REGION Network 29: Encoder Wals Function Block
   RUNG wire#powerrail
      "FB_EncoderFeedback_Aanvoerband"(CounterTag := "EncoderBand_RawCounter", Position_Offset := "PositionManagement".Axis_1.Values."Position Offset", Pulsfactor := "PositionManagement".Axis_1.Values.Pulsfactor, Position_Correction := "PositionManagement".Axis_1.Values."Axis Correction", ReferenceRun_Command := "PositionManagement".Axis_1.Commands."Start Ref Run", ReferenceSwitch := "Zpuls_Encoder_Band", ReferencePosition := "PositionManagement".Axis_1.Values."Reference Position", Scaled_Position => #Axis1_ScaledPosition, Actual_Enc_Pos => #Axis1_ActualEncPosition, AxisDB_Connection => "PositionManagement".Data.Actual_Axis1_Position)
   END_RUNG
   // the same network as SCL:
   "FB_EncoderFeedback_Aanvoerband"(CounterTag := "EncoderBand_RawCounter",   // "FB_EncoderFeedback"
                           Position_Offset := "PositionManagement".Axis_1.Values."Position Offset",
                           Pulsfactor := "PositionManagement".Axis_1.Values.Pulsfactor,
                           Position_Correction := "PositionManagement".Axis_1.Values."Axis Correction",
                           ReferenceRun_Command := "PositionManagement".Axis_1.Commands."Start Ref Run",
                           ReferenceSwitch := "Zpuls_Encoder_Band",
                           ReferencePosition := "PositionManagement".Axis_1.Values."Reference Position",
                           Scaled_Position => #Axis1_ScaledPosition,
                           Actual_Enc_Pos => #Axis1_ActualEncPosition,
                           AxisDB_Connection => "PositionManagement".Data.Actual_Axis1_Position);
END_REGION

REGION Network 30: SystemTime
   "PLCMemory".SystemTime := TIME_TCK();
END_REGION
END_ORGANIZATION_BLOCK

// folder: Blocks

FUNCTION_BLOCK "ESB_Flash_Warning_Block"   // FB1, FBD
{ S7_Optimized_Access := 'FALSE' }
VERSION : 0.1
   VAR_INPUT
      "Safety Feedback Contact" : Bool;
      "WarningTimer Time 1" : Time := T#150ms;
      "WarningTimer Time 2" : Time := T#150ms;
   END_VAR
   VAR_OUTPUT
      "Warning Ouput Contact" : Bool;
      "ET WarningTimer 1" : Time;
      "ET WarningTimer 2" : Time;
   END_VAR
   VAR_TEMP
      SafetyTakeoverContact : Bool;
   END_VAR
   VAR_TEMP   // added for the SCL form of the ladder/FBD networks
      _w1 : Bool;
   END_VAR
BEGIN

REGION Network 1: Flash Warning
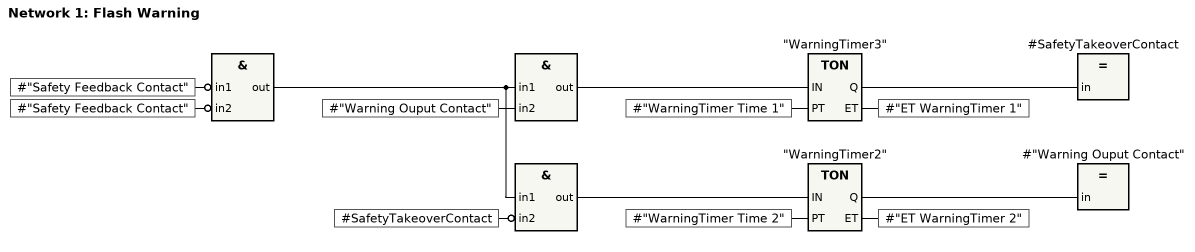
   #_w1 := NOT #"Safety Feedback Contact" AND NOT #"Safety Feedback Contact";
   "WarningTimer3".TON(IN := #_w1 AND #"Warning Ouput Contact",
                       PT := #"WarningTimer Time 1",
                       ET => #"ET WarningTimer 1");
   #SafetyTakeoverContact := "WarningTimer3".Q;
   "WarningTimer2".TON(IN := #_w1 AND NOT #SafetyTakeoverContact,
                       PT := #"WarningTimer Time 2",
                       ET => #"ET WarningTimer 2");
   #"Warning Ouput Contact" := "WarningTimer2".Q;
END_REGION
END_FUNCTION_BLOCK

FUNCTION_BLOCK "Delayed_Message_Function"   // FB2, FBD
TITLE = Delayed Message Function
{ S7_Optimized_Access := 'FALSE' }
VERSION : 0.1
// Functionblock For Delaying Message Function for example for filling an magazine or waiting for an signal. It is possible to adjust Time with the Dleay Time Message Input. The FlashTimer Time 1 & 2 ar for adjusting the flashing time of the ouput LED.
   VAR_INPUT
      "Override Message" : Bool;
      "Sensor Input 1" : Bool;
      "Sensor Input 2" : Bool := true;
      "Delay Time Message" : Time := T#1S_500MS;
      "FlashTimer Time 1" : Time := T#200ms;
      "FlashTimer Time 2" : Time := T#200ms;
   END_VAR
   VAR_OUTPUT
      "Output Signal" : Bool;
      "Output Signal Halt" : Bool;
      "ET Delayed Timer" : Time;
      "Output LED Flashing" : Bool;
   END_VAR
   VAR_TEMP
      "Internal Delayed Signal" : Bool;
   END_VAR
   VAR_TEMP   // added for the SCL form of the ladder/FBD networks
      _w1 : Bool;
   END_VAR
BEGIN

REGION Network 1: Delayed Signal to Outputs
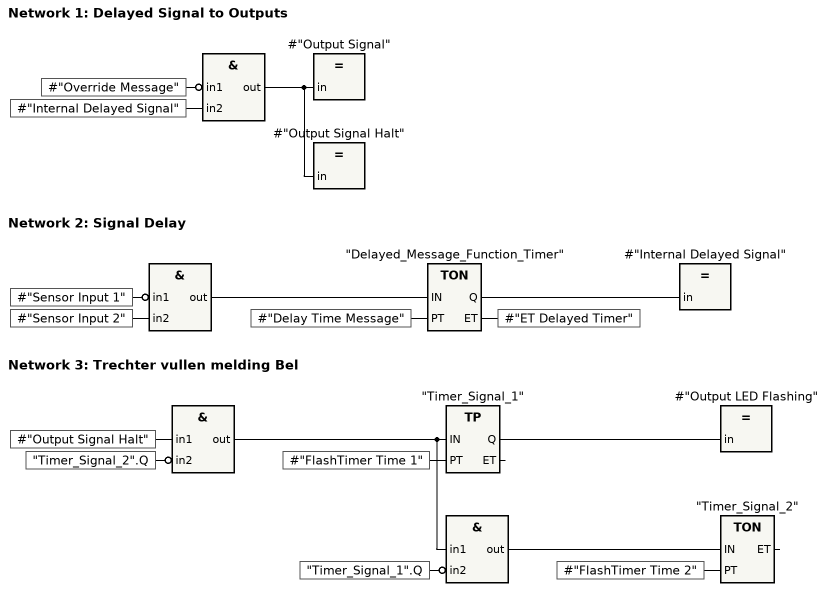
   #"Output Signal" := NOT #"Override Message" AND #"Internal Delayed Signal";
   #"Output Signal Halt" := #"Output Signal";
END_REGION

REGION Network 2: Signal Delay
   "Delayed_Message_Function_Timer".TON(IN := NOT #"Sensor Input 1" AND #"Sensor Input 2",
                           PT := #"Delay Time Message",
                           ET => #"ET Delayed Timer");
   #"Internal Delayed Signal" := "Delayed_Message_Function_Timer".Q;
END_REGION

REGION Network 3: Trechter vullen melding Bel
   #_w1 := #"Output Signal Halt" AND NOT "Timer_Signal_2".Q;
   "Timer_Signal_1".TP(IN := #_w1, PT := #"FlashTimer Time 1");
   #"Output LED Flashing" := "Timer_Signal_1".Q;
   "Timer_Signal_2".TON(IN := #_w1 AND NOT "Timer_Signal_1".Q, PT := #"FlashTimer Time 2");
END_REGION
END_FUNCTION_BLOCK

FUNCTION_BLOCK "Alarm_Axis_Position_Function"   // FB3, FBD
TITLE = Alarm Axis not in Position
{ S7_Optimized_Access := 'FALSE' }
VERSION : 0.1
   VAR_INPUT
      "Axis FWD command" : Bool;
      "Axis Feedback (Sensor) signal" : Bool;
      "Axis Encoder Singal" : Real;
      "Axis Command Position" : Real;
      "Sensor Controlled (HIGH) - Position Controlled (LOW)" : Bool;
      "CheckTime Setting" : Time := T#5S;
   END_VAR
   VAR_OUTPUT
      "Alarm BOOL" : Bool;
      "Alarm WORD" : Bool;
   END_VAR
   VAR_TEMP
      "Axis Feedback Internal" : Bool;
      "Axis Encoder On Position" : Bool;
      "Axis Sensor On Position" : Bool;
      "Axis Measuring Mode" : Bool;
   END_VAR
BEGIN

REGION Network 1: When axis is spinning start timer
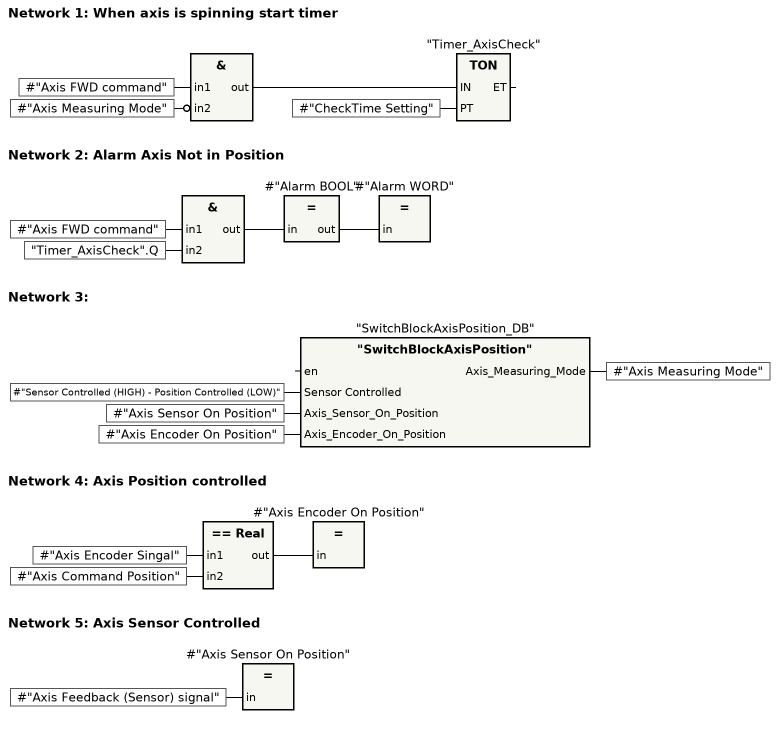
   "Timer_AxisCheck".TON(IN := #"Axis FWD command" AND NOT #"Axis Measuring Mode", PT := #"CheckTime Setting");
END_REGION

REGION Network 2: Alarm Axis Not in Position
   #"Alarm BOOL" := #"Axis FWD command" AND "Timer_AxisCheck".Q;
   #"Alarm WORD" := #"Alarm BOOL";
END_REGION

REGION Network 3
   "SwitchBlockAxisPosition_DB"("Sensor Controlled" := #"Sensor Controlled (HIGH) - Position Controlled (LOW)",   // "SwitchBlockAxisPosition"
                           Axis_Sensor_On_Position := #"Axis Sensor On Position",
                           Axis_Encoder_On_Position := #"Axis Encoder On Position",
                           Axis_Measuring_Mode => #"Axis Measuring Mode");
END_REGION

REGION Network 4: Axis Position controlled
   #"Axis Encoder On Position" := #"Axis Encoder Singal" = #"Axis Command Position";
END_REGION

REGION Network 5: Axis Sensor Controlled
   #"Axis Sensor On Position" := #"Axis Feedback (Sensor) signal";
END_REGION
END_FUNCTION_BLOCK

FUNCTION_BLOCK "SwitchBlockAxisPosition"   // FB4, SCL
{ S7_Optimized_Access := 'FALSE' }
VERSION : 0.1
   VAR_INPUT
      "Sensor Controlled" : Bool;
      Axis_Sensor_On_Position : Bool;
      Axis_Encoder_On_Position : Bool;
   END_VAR
   VAR_OUTPUT
      Axis_Measuring_Mode : Bool;
   END_VAR
BEGIN
   IF #"Sensor Controlled" THEN
       #Axis_Measuring_Mode := #Axis_Sensor_On_Position;
   ELSE
       #Axis_Measuring_Mode := #Axis_Encoder_On_Position;
   END_IF;
END_FUNCTION_BLOCK

FUNCTION_BLOCK "DriveConfirmation_Function"   // FB5, FBD
TITLE = Drive Confirmation Function Block
{ S7_Optimized_Access := 'FALSE' }
VERSION : 0.1
   VAR_INPUT
      "System RUN" : Bool;
      "Drive Ouput Q" : Bool;
      "Drive Ready Signal" : Bool;
      DelayTime : Time := T#1s;
   END_VAR
   VAR_OUTPUT
      "Timer ET" : Time;
      "Ouput WORD" : Bool;
   END_VAR
BEGIN

REGION Network 1: Confirmation Drive
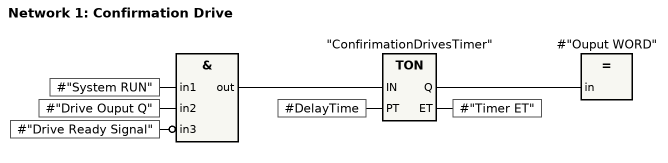
   "ConfirimationDrivesTimer".TON(IN := #"System RUN" AND #"Drive Ouput Q" AND NOT #"Drive Ready Signal",
                           PT := #DelayTime,
                           ET => #"Timer ET");
   #"Ouput WORD" := "ConfirimationDrivesTimer".Q;
END_REGION
END_FUNCTION_BLOCK

FUNCTION_BLOCK "2in-1out_Block"   // FB6, FBD
{ S7_Optimized_Access := 'FALSE' }
VERSION : 0.1
   VAR_INPUT
      "Input Contact 1" : Bool;
      "Input Contact 2" : Bool;
   END_VAR
   VAR_OUTPUT
      "Output Contact 1" : Bool;
   END_VAR
BEGIN

REGION Network 1: Network Default
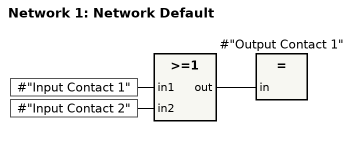
   #"Output Contact 1" := #"Input Contact 1" OR #"Input Contact 2";
END_REGION
END_FUNCTION_BLOCK

FUNCTION_BLOCK "Override_Block_Safety"   // FB7, FBD
TITLE = Override Block Safety.
{ S7_Optimized_Access := 'FALSE' }
VERSION : 0.1
   VAR_INPUT
      "SAFE Q 1" : Bool;
      "SAFE Q 2" : Bool;
      "Override Contact" : Bool;
      "Delay Timer" : Time;
   END_VAR
   VAR_OUTPUT
      "SAFE Output Contact" : Bool;
      "Timer ET" : Time;
   END_VAR
BEGIN

REGION Network 1: SAFETY - OVERRIDE
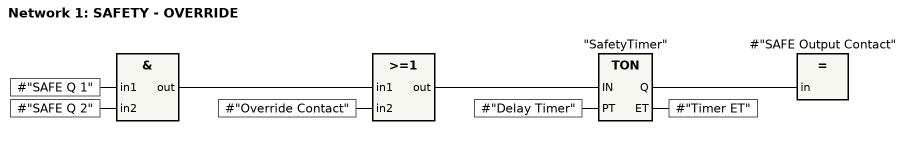
   "SafetyTimer".TON(IN := (#"SAFE Q 1" AND #"SAFE Q 2") OR #"Override Contact",
                     PT := #"Delay Timer",
                     ET => #"Timer ET");
   #"SAFE Output Contact" := "SafetyTimer".Q;
END_REGION
END_FUNCTION_BLOCK

FUNCTION_BLOCK "Ouput_Function_1"   // FB8, FBD
TITLE = Ouput Controller Function Block
{ S7_Optimized_Access := 'FALSE' }
VERSION : 0.1
   VAR_INPUT
      "Stop Contact" : Bool;
      "Manual Command" : Bool;
      "Auto Command" : Bool;
      "Option Command" : Bool;
      "Disable Command" : Bool;
   END_VAR
   VAR_OUTPUT
      "Ouput Signal" : Bool;
   END_VAR
BEGIN

REGION Network 1: Ouput Controller
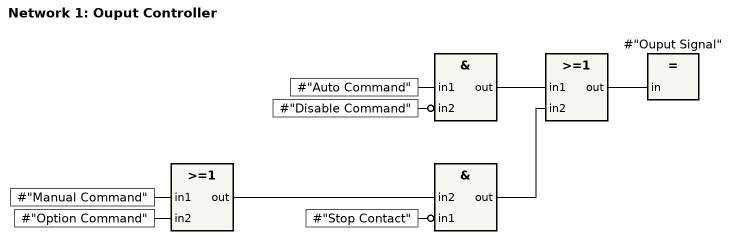
   #"Ouput Signal" := (#"Auto Command" AND NOT #"Disable Command") OR ((#"Manual Command" OR #"Option Command") AND NOT #"Stop Contact");
END_REGION
END_FUNCTION_BLOCK

FUNCTION_BLOCK "ResetOuputs_Function"   // FB9, LAD
TITLE = Reset Ouput Functions With Commands
{ S7_Optimized_Access := 'FALSE' }
VERSION : 0.1
   VAR_INPUT
      StopCommand_NC : Bool;
      StopCommand_NO : Bool;
   END_VAR
   VAR_OUTPUT
      Output_1 : Bool;
      Output_2 : Bool;
      Output_3 : Bool;
      Output_4 : Bool;
      Output_5 : Bool;
      Output_6 : Bool;
      Output_7 : Bool;
      Output_8 : Bool;
      Output_9 : Bool;
      Output_10 : Bool;
   END_VAR
BEGIN

REGION Network 1: NW1
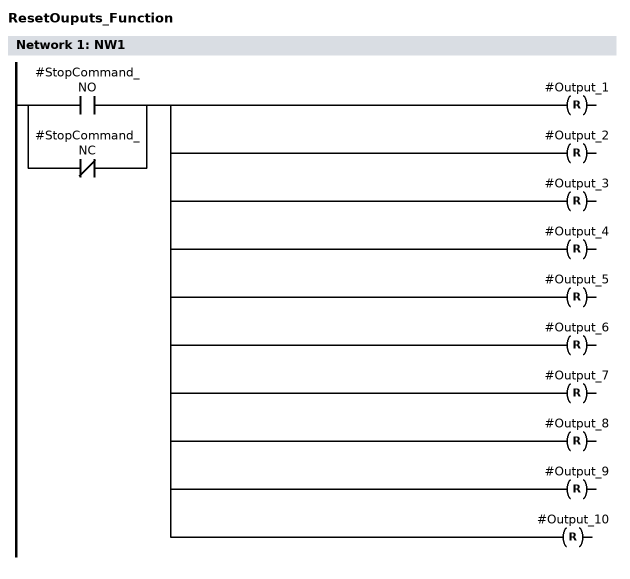
   RUNG wire#powerrail
      Contact( #StopCommand_NO )
      wire#w1
      R_Coil( #Output_1 )
   END_RUNG
   RUNG wire#powerrail
      I_Contact( #StopCommand_NC )
   END_RUNG wire#w1
   RUNG wire#w1
      R_Coil( #Output_2 )
   END_RUNG
   RUNG wire#w1
      R_Coil( #Output_3 )
   END_RUNG
   RUNG wire#w1
      R_Coil( #Output_4 )
   END_RUNG
   RUNG wire#w1
      R_Coil( #Output_5 )
   END_RUNG
   RUNG wire#w1
      R_Coil( #Output_6 )
   END_RUNG
   RUNG wire#w1
      R_Coil( #Output_7 )
   END_RUNG
   RUNG wire#w1
      R_Coil( #Output_8 )
   END_RUNG
   RUNG wire#w1
      R_Coil( #Output_9 )
   END_RUNG
   RUNG wire#w1
      R_Coil( #Output_10 )
   END_RUNG
   // the same network as SCL:
   IF #StopCommand_NO OR NOT #StopCommand_NC THEN
       #Output_1 := FALSE;
       #Output_2 := FALSE;
       #Output_3 := FALSE;
       #Output_4 := FALSE;
       #Output_5 := FALSE;
       #Output_6 := FALSE;
       #Output_7 := FALSE;
       #Output_8 := FALSE;
       #Output_9 := FALSE;
       #Output_10 := FALSE;
   END_IF;
END_REGION
END_FUNCTION_BLOCK

FUNCTION_BLOCK "Blinker"   // FB15, SCL
{ S7_Optimized_Access := 'FALSE' }
VERSION : 0.1
   VAR_INPUT
      Enable : Bool;
      BlinkTime : Time := T#500ms;
   END_VAR
   VAR_OUTPUT
      Q_Blink : Bool;
      Q_Blink2 : Bool;
   END_VAR
   VAR
      BlinkTimer : TON;
   END_VAR
   VAR_TEMP
      LastToggleTime : Time;
   END_VAR
BEGIN
   // Logica
   IF #Enable THEN
       #BlinkTimer(IN := TRUE,
                   PT := #BlinkTime);   // Correct gebruik van PT

       IF #BlinkTimer.Q THEN
           #Q_Blink := NOT #Q_Blink;                // Toggle uitgang
           #Q_Blink2 := NOT #Q_Blink2;
           #BlinkTimer(IN := FALSE,
                       PT := #BlinkTime); // Reset timer (verplicht opnieuw PT meegeven)
       END_IF;

   ELSE
       #BlinkTimer(IN := FALSE,
                   PT := #BlinkTime);  // Timer uitzetten
       #Q_Blink := FALSE; // Uitgang terug laag
       #Q_Blink2 := FALSE;
   END_IF;
END_FUNCTION_BLOCK

FUNCTION_BLOCK "BlowOff_Timer"   // FB16, SCL
{ S7_Optimized_Access := 'FALSE' }
VERSION : 0.1
   VAR_INPUT
      Enable : Bool;
      CycleTime : Time;
      PulseDuration : Time;
      NowTime : Time;
   END_VAR
   VAR_OUTPUT
      Q_Pulse : Bool;
   END_VAR
   VAR
      CycleTimer : TON;
      PulseTimer : TON;
      State : Int;
      S_PEXT : Int;
   END_VAR
   VAR_TEMP
      PulseActive : Bool;
      StartPulse : Bool;
      TriggerPulse : Bool;
      PulseBusy : Bool;
      DummyWord : Word;
      DummyWord2 : Bool;
      T1 : Int;
      PulseStartTime : Time;
      LastPulseEndTime : Time;
      LastPulseTime : Time;
   END_VAR
BEGIN
   // Logica
   IF #Enable THEN
       // Start cyclische timer
       #CycleTimer(IN := TRUE,
                   PT := #CycleTime);

       IF #CycleTimer.Q THEN
           // Start puls-timer als cyclus voorbij is
           #PulseTimer(IN := TRUE,
                       PT := #PulseDuration);

           // Reset de CycleTimer voor de volgende cyclus
           #CycleTimer(IN := FALSE,
                       PT := #CycleTime);
       END_IF;

       // Puls-timer logica
       IF #PulseTimer.IN THEN
           #Q_Pulse := TRUE;

           IF #PulseTimer.Q THEN
               // Puls voorbij, pulse output uit
               #PulseTimer(IN := FALSE,
                           PT := #PulseDuration);
               #Q_Pulse := FALSE;
           END_IF;
       ELSE
           #Q_Pulse := FALSE;
       END_IF;

   ELSE
       // Alles resetten bij disable
       #CycleTimer(IN := FALSE,
                   PT := #CycleTime);
       #PulseTimer(IN := FALSE,
                   PT := #PulseDuration);
       #Q_Pulse := FALSE;
   END_IF;
END_FUNCTION_BLOCK

FUNCTION_BLOCK "ProductBuffer"   // FB17, SCL
{ S7_Optimized_Access := 'FALSE' }
VERSION : 0.1
   VAR_INPUT
      SensorInput : Bool;
      TimeDelay : Time;
      TriggerFeedback : Bool;
   END_VAR
   VAR_OUTPUT
      TriggerMovement : Bool;
      ProductCount : Int;
   END_VAR
   VAR
      PrevSensor : Bool;
      DelayTimer : TON;
      MovementActive : Bool;
   END_VAR
BEGIN
   // Flankdetectie op sensor
   IF #SensorInput AND NOT #PrevSensor THEN
       IF #ProductCount < 32767 THEN
           #ProductCount := #ProductCount + 1;
       END_IF;
   END_IF;
   #PrevSensor := #SensorInput;

   // Timer mag alleen lopen als:
   // - Er producten zijn
   // - Er geen beweging actief is
   IF (#ProductCount > 0) AND (NOT #MovementActive) THEN
       #DelayTimer(IN := TRUE,
                   PT := #TimeDelay);
   ELSE
       #DelayTimer(IN := FALSE,
                   PT := #TimeDelay);
   END_IF;

   // Als de timer klaar is → activeer beweging en zet MovementActive
   IF #DelayTimer.Q THEN
       #TriggerMovement := TRUE;
       #MovementActive := TRUE;
       #ProductCount := #ProductCount - 1;
       #DelayTimer(IN := FALSE,
                   PT := #TimeDelay); // Reset timer
   END_IF;

   // Wacht op TriggerFeedback om TriggerMovement terug laag te zetten
   IF #MovementActive AND #TriggerFeedback THEN
       #TriggerMovement := FALSE;
       #MovementActive := FALSE;
   END_IF;
END_FUNCTION_BLOCK

FUNCTION_BLOCK "ProductBuffer_V2"   // FB18, SCL
{ S7_Optimized_Access := 'FALSE' }
VERSION : 0.1
   VAR_INPUT
      SensorInput : Bool;
      SensorManual : Bool;
      TimeDelay : Time;
      SystemTime : Time;
      TriggerFeedback : Bool;
   END_VAR
   VAR_OUTPUT
      TriggerMovement : Bool;
      InsertIndex : Int;
      ProductCount : Int;
      SystemTicks : DInt;
   END_VAR
   VAR
      ProductQueue : Array[0..1] of "ProductEntry";
      StartTimes : Struct
         _0 : Time;
         _1 : Time;
         _2 : Time;
         _3 : Time;
         _4 : Time;
         _5 : Time;
         _6 : Time;
         _7 : Time;
         _8 : Time;
         _9 : Time;
      END_STRUCT;
      Actives : Struct
         _0 : Bool;
         _1 : Bool;
         _2 : Bool;
         _3 : Bool;
         _4 : Bool;
         _5 : Bool;
         _6 : Bool;
         _7 : Bool;
         _8 : Bool;
         _9 : Bool;
      END_STRUCT;
      PrevSensor : Bool;
      MovementActive : Bool;
      i : Int;
      Elapsed : DInt;
   END_VAR
BEGIN
   // Flankdetectie sensor
   IF #SensorInput AND NOT #PrevSensor THEN
       CASE #InsertIndex MOD 10 OF
           0:
               IF NOT #Actives._0 THEN
                   #Actives._0 := TRUE;
                   #StartTimes._0 := #SystemTime;
               END_IF;
           1:
               IF NOT #Actives._1 THEN
                   #Actives._1 := TRUE;
                   #StartTimes._1 := #SystemTime;
               END_IF;
           2:
               IF NOT #Actives._2 THEN
                   #Actives._2 := TRUE;
                   #StartTimes._2 := #SystemTime;
               END_IF;
           3:
               IF NOT #Actives._3 THEN
                   #Actives._3 := TRUE;
                   #StartTimes._3 := #SystemTime;
               END_IF;
           4:
               IF NOT #Actives._4 THEN
                   #Actives._4 := TRUE;
                   #StartTimes._4 := #SystemTime;
               END_IF;
           5:
               IF NOT #Actives._5 THEN
                   #Actives._5 := TRUE;
                   #StartTimes._5 := #SystemTime;
               END_IF;
           6:
               IF NOT #Actives._6 THEN
                   #Actives._6 := TRUE;
                   #StartTimes._6 := #SystemTime;
               END_IF;
           7:
               IF NOT #Actives._7 THEN
                   #Actives._7 := TRUE;
                   #StartTimes._7 := #SystemTime;
               END_IF;
           8:
               IF NOT #Actives._8 THEN
                   #Actives._8 := TRUE;
                   #StartTimes._8 := #SystemTime;
               END_IF;
           9:
               IF NOT #Actives._9 THEN
                   #Actives._9 := TRUE;
                   #StartTimes._9 := #SystemTime;
               END_IF;
       END_CASE;
       #InsertIndex := (#InsertIndex + 1) MOD 10;
   END_IF;

   #PrevSensor := #SensorInput;

   // Tellen hoeveel producten actief zijn
   #ProductCount := 0;
   IF #Actives._0 THEN
       #ProductCount := #ProductCount + 1;
   END_IF;
   IF #Actives._1 THEN
       #ProductCount := #ProductCount + 1;
   END_IF;
   IF #Actives._2 THEN
       #ProductCount := #ProductCount + 1;
   END_IF;
   IF #Actives._3 THEN
       #ProductCount := #ProductCount + 1;
   END_IF;
   IF #Actives._4 THEN
       #ProductCount := #ProductCount + 1;
   END_IF;
   IF #Actives._5 THEN
       #ProductCount := #ProductCount + 1;
   END_IF;
   IF #Actives._6 THEN
       #ProductCount := #ProductCount + 1;
   END_IF;
   IF #Actives._7 THEN
       #ProductCount := #ProductCount + 1;
   END_IF;
   IF #Actives._8 THEN
       #ProductCount := #ProductCount + 1;
   END_IF;
   IF #Actives._9 THEN
       #ProductCount := #ProductCount + 1;
   END_IF;

   // Beweging starten als een product klaar is en geen andere beweging actief is
   IF NOT #MovementActive THEN
       IF #Actives._0 THEN
           #Elapsed := TIME_TO_DINT(#SystemTime) - TIME_TO_DINT(#StartTimes._0);
           IF #Elapsed >= TIME_TO_DINT(#TimeDelay) THEN
               #TriggerMovement := TRUE;
               #MovementActive := TRUE;
               #Actives._0 := FALSE;
           END_IF;
       ELSIF #Actives._1 THEN
           #Elapsed := TIME_TO_DINT(#SystemTime) - TIME_TO_DINT(#StartTimes._1);
           IF #Elapsed >= TIME_TO_DINT(#TimeDelay) THEN
               #TriggerMovement := TRUE;
               #MovementActive := TRUE;
               #Actives._1 := FALSE;
           END_IF;
       ELSIF #Actives._2 THEN
           #Elapsed := TIME_TO_DINT(#SystemTime) - TIME_TO_DINT(#StartTimes._2);
           IF #Elapsed >= TIME_TO_DINT(#TimeDelay) THEN
               #TriggerMovement := TRUE;
               #MovementActive := TRUE;
               #Actives._2 := FALSE;
           END_IF;
       ELSIF #Actives._3 THEN
           #Elapsed := TIME_TO_DINT(#SystemTime) - TIME_TO_DINT(#StartTimes._3);
           IF #Elapsed >= TIME_TO_DINT(#TimeDelay) THEN
               #TriggerMovement := TRUE;
               #MovementActive := TRUE;
               #Actives._3 := FALSE;
           END_IF;
       ELSIF #Actives._4 THEN
           #Elapsed := TIME_TO_DINT(#SystemTime) - TIME_TO_DINT(#StartTimes._4);
           IF #Elapsed >= TIME_TO_DINT(#TimeDelay) THEN
               #TriggerMovement := TRUE;
               #MovementActive := TRUE;
               #Actives._4 := FALSE;
           END_IF;
       ELSIF #Actives._5 THEN
           #Elapsed := TIME_TO_DINT(#SystemTime) - TIME_TO_DINT(#StartTimes._5);
           IF #Elapsed >= TIME_TO_DINT(#TimeDelay) THEN
               #TriggerMovement := TRUE;
               #MovementActive := TRUE;
               #Actives._5 := FALSE;
           END_IF;
       ELSIF #Actives._6 THEN
           #Elapsed := TIME_TO_DINT(#SystemTime) - TIME_TO_DINT(#StartTimes._6);
           IF #Elapsed >= TIME_TO_DINT(#TimeDelay) THEN
               #TriggerMovement := TRUE;
               #MovementActive := TRUE;
               #Actives._6 := FALSE;
           END_IF;
       ELSIF #Actives._7 THEN
           #Elapsed := TIME_TO_DINT(#SystemTime) - TIME_TO_DINT(#StartTimes._7);
           IF #Elapsed >= TIME_TO_DINT(#TimeDelay) THEN
               #TriggerMovement := TRUE;
               #MovementActive := TRUE;
               #Actives._7 := FALSE;
           END_IF;
       ELSIF #Actives._8 THEN
           #Elapsed := TIME_TO_DINT(#SystemTime) - TIME_TO_DINT(#StartTimes._8);
           IF #Elapsed >= TIME_TO_DINT(#TimeDelay) THEN
               #TriggerMovement := TRUE;
               #MovementActive := TRUE;
               #Actives._8 := FALSE;
           END_IF;
       ELSIF #Actives._9 THEN
           #Elapsed := TIME_TO_DINT(#SystemTime) - TIME_TO_DINT(#StartTimes._9);
           IF #Elapsed >= TIME_TO_DINT(#TimeDelay) THEN
               #TriggerMovement := TRUE;
               #MovementActive := TRUE;
               #Actives._9 := FALSE;
           END_IF;
       END_IF;
   END_IF;

   // Beweging beëindigen na feedback
   IF #MovementActive AND #TriggerFeedback THEN
       #TriggerMovement := FALSE;
       #MovementActive := FALSE;
   END_IF;
END_FUNCTION_BLOCK

FUNCTION "SCL_Block" : Void   // FC10, SCL
{ S7_Optimized_Access := 'FALSE' }
VERSION : 0.1
BEGIN
   // Reset de Word variabelen aan het begin van elke cyclus
   "Alarms".AlarmsWord := 0;
   "Alarms".HMI_Alarm_Drive1 := 0;
   "Alarms".HMI_Alarm_Drive2 := 0;
   "Alarms".HMI_Alarm_Drive3 := 0;
   "Alarms".HMI_Alarm_Drive4 := 0;
   "Alarms".HMI_Alarm_Drive5 := 0;

   // Controleer de alarmen en zet de respectievelijke bits aan
   IF "Alarms".AlarmStruct.Alarm_Product_Not_Position THEN
       "Alarms".AlarmsWord := "Alarms".AlarmsWord OR WORD#1; // Zet bit 0 aan
   END_IF;

   IF "Alarms".AlarmStruct.Alarm_Axis_Not_Position THEN
       "Alarms".AlarmsWord := "Alarms".AlarmsWord OR WORD#2; // Zet bit 1 aan
   END_IF;

   IF "Alarms".AlarmStruct.Alarm_Drive1 THEN
       "Alarms".HMI_Alarm_Drive1 := "Alarms".HMI_Alarm_Drive1 OR WORD#1; // Zet bit 2 aan
   END_IF;

   IF "Alarms".AlarmStruct.Alarm_Drive2 THEN
       "Alarms".HMI_Alarm_Drive2 := "Alarms".HMI_Alarm_Drive2 OR WORD#1; // Zet bit 3 aan
   END_IF;

   IF "Alarms".AlarmStruct.Alarm_Drive3 THEN
       "Alarms".HMI_Alarm_Drive3 := "Alarms".HMI_Alarm_Drive3 OR WORD#1; // Zet bit 4 aan
   END_IF;

   IF "Alarms".AlarmStruct.Alarm_Drive4 THEN
       "Alarms".HMI_Alarm_Drive4 := "Alarms".HMI_Alarm_Drive4 OR WORD#1; // Zet bit 5 aan
   END_IF;

   IF "Alarms".AlarmStruct.Alarm_Drive5 THEN
       "Alarms".HMI_Alarm_Drive5 := "Alarms".HMI_Alarm_Drive5 OR WORD#1; // Zet bit 6 aan
   END_IF;


   // Position Program Axis 3 (Wals)

   // Configureer de timer om elke 0,5 seconde af te lopen
   "Timer_0_5s".TON(IN := TRUE,
   PT := "PLCMemory"."Encoder PulsOffset");

   // Controleer of de timer is afgelopen
   IF "Timer_0_5s".Q THEN
       // Verhoog of verlaag de positie afhankelijk van de aandrijfsignalen
       IF "Drive 3 RUN FWD" THEN
           "PLCMemory".EncoderPosition := "PLCMemory".EncoderPosition + "PLCMemory".StepSize; // Verhoog met de stepgrootte
       ELSIF "Drive 3 REV" THEN
           "PLCMemory".EncoderPosition := "PLCMemory".EncoderPosition - "PLCMemory".StepSize; // Verlaag met de stepgrootte
       END_IF;

       // Wrapping van de positie bij overschrijden van 360 graden of onder 0 graden
       IF "PLCMemory".EncoderPosition >= 360.0 THEN
           "PLCMemory".EncoderPosition := 0.0;  // Wrapping naar 0 als de positie 360 overschrijdt
       ELSIF "PLCMemory".EncoderPosition < 0.0 THEN
           "PLCMemory".EncoderPosition := 360.0; // Wrapping naar 360 als de positie onder 0 gaat
       END_IF;

       // Reset de timer
       "Timer_0_5s".TON (IN := FALSE,
                         PT := "PLCMemory"."Encoder PulsOffset"); // Reset de timer zodat deze opnieuw kan starten
   END_IF;

   // Homing logica
   IF "Sensor Wals (Option)" THEN
       "PLCMemory".EncoderPosition := 0.0;  // Reset de positie naar 0 als de sensor wordt geactiveerd
   END_IF;



   //Drive Servo Control Here:
   /// Desired Position Axis 3

   // Controleer of de HMI-knop is ingedrukt en er een gewenste positie is ingesteld
   //IF "HMI_Des_Pos_Axis3" THEN
       //"GoButtonPressed" := TRUE; // HMI-knop is ingedrukt, start beweging
   //END_IF;

   // Beveiliging voor de Desired_Encoder_Position: Zorg dat de waarde tussen 0 en 360 blijft
   //IF "PLCMemory".Desired_Encoder_Position > 360.0 THEN
     //  "PLCMemory".Desired_Encoder_Position := 360.0;  // Zet naar 360 als de waarde boven 360 ligt
   //ELSIF "PLCMemory".Desired_Encoder_Position < 0.0 THEN
       //"PLCMemory".Desired_Encoder_Position := 0.0;  // Zet naar 0 als de waarde onder 0 ligt
   //END_IF;

   // Wrapping van de gewenste positie: Als de gewenste positie 360 is, zet deze dan op 0
   //IF "PLCMemory".Desired_Encoder_Position = 360.0 THEN
      // "PLCMemory".Desired_Encoder_Position := 0.0;  // Wrapping naar 0 als de gewenste positie 360 is
   //END_IF;

   // Voer beweging uit totdat de gewenste positie is bereikt
   //IF "GoButtonPressed" THEN
       // Bepaal de bewegingsrichting en start de beweging
     //  IF "PLCMemory".EncoderPosition < "PLCMemory".Desired_Encoder_Position - "PLCMemory".Tolerance THEN
           // Beweeg vooruit met StepSize als snelheid
         //  "PLCMemory".EncoderPosition := "PLCMemory".EncoderPosition + "PLCMemory".StepSize;
        //   "Drive_3_Manual" := TRUE;   // Activeer vooruitbeweging
         //  "Drive 3 REV" := FALSE;     // Zorg dat achteruitbeweging uit is

     //  ELSIF "PLCMemory".EncoderPosition > "PLCMemory".Desired_Encoder_Position + "PLCMemory".Tolerance THEN
           // Beweeg achteruit met StepSize als snelheid
        //   "PLCMemory".EncoderPosition := "PLCMemory".EncoderPosition - "PLCMemory".StepSize;
       //    "Drive_3_Manual" := FALSE;  // Zorg dat vooruitbeweging uit is
       //    "Drive 3 REV" := TRUE;      // Activeer achteruitbeweging

      // ELSE
           // Stop de beweging zodra de positie binnen de tolerantie komt
         //  "Drive_3_Manual" := FALSE;    // Zet vooruitbeweging uit
        //   "Drive 3 REV" := FALSE;       // Zet achteruitbeweging uit
        //   "GoButtonPressed" := FALSE;   // Zet de Go-knop uit om verdere beweging te stoppen
      // END_IF;
   //END_IF;
END_FUNCTION

FUNCTION "SafetyFunction_Block" : Void   // FC12, LAD
{ S7_Optimized_Access := 'FALSE' }
VERSION : 0.1
   VAR_INPUT
      "ESB NC Contact" : Bool;
      "ESB NO Contact" : Bool;
      "Reset NO Contact" : Bool;
      "SAFE door 1 NC Contact" : Bool;
      "SAFE door 2 NC Contact" : Bool;
      "Safety Relais NO Contact" : Bool;
   END_VAR
   VAR_OUTPUT
      SAFE_OK_Signal : Bool;
   END_VAR
BEGIN

REGION Network 1: +MC-21K6:1 - Noodstop Circuit
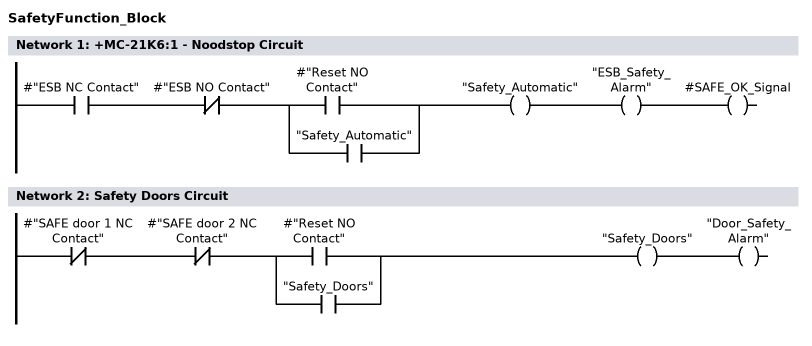
   RUNG wire#powerrail
      Contact( #"ESB NC Contact" )
      I_Contact( #"ESB NO Contact" )
      wire#w1
      Contact( #"Reset NO Contact" )
      wire#w2
      Coil( "Safety_Automatic" )
      Coil( "ESB_Safety_Alarm" )
      Coil( #SAFE_OK_Signal )
   END_RUNG
   RUNG wire#w1
      Contact( "Safety_Automatic" )
   END_RUNG wire#w2
   // the same network as SCL:
   "Safety_Automatic" := #"ESB NC Contact" AND NOT #"ESB NO Contact" AND (#"Reset NO Contact" OR "Safety_Automatic");
   "ESB_Safety_Alarm" := "Safety_Automatic";
   #SAFE_OK_Signal := "Safety_Automatic";
END_REGION

REGION Network 2: Safety Doors Circuit
   RUNG wire#powerrail
      I_Contact( #"SAFE door 1 NC Contact" )
      I_Contact( #"SAFE door 2 NC Contact" )
      wire#w1
      Contact( #"Reset NO Contact" )
      wire#w2
      Coil( "Safety_Doors" )
      Coil( "Door_Safety_Alarm" )
   END_RUNG
   RUNG wire#w1
      Contact( "Safety_Doors" )
   END_RUNG wire#w2
   // the same network as SCL:
   "Safety_Doors" := NOT #"SAFE door 1 NC Contact" AND NOT #"SAFE door 2 NC Contact" AND (#"Reset NO Contact" OR "Safety_Doors");
   "Door_Safety_Alarm" := "Safety_Doors";
END_REGION
END_FUNCTION

FUNCTION "SystemRUN_Block" : Void   // FC13, LAD
{ S7_Optimized_Access := 'FALSE' }
VERSION : 0.1
   VAR_INPUT
      "Safety Relais Contact" : Bool;
      "Stop Machine NC Contact" : Bool;
      "Fill Magzine Contact" : Bool;
      "Start Machine NO Contact" : Bool;
   END_VAR
   VAR_OUTPUT
      "Run Output Lamp" : Bool;
   END_VAR
BEGIN

REGION Network 1: Systeem RUN
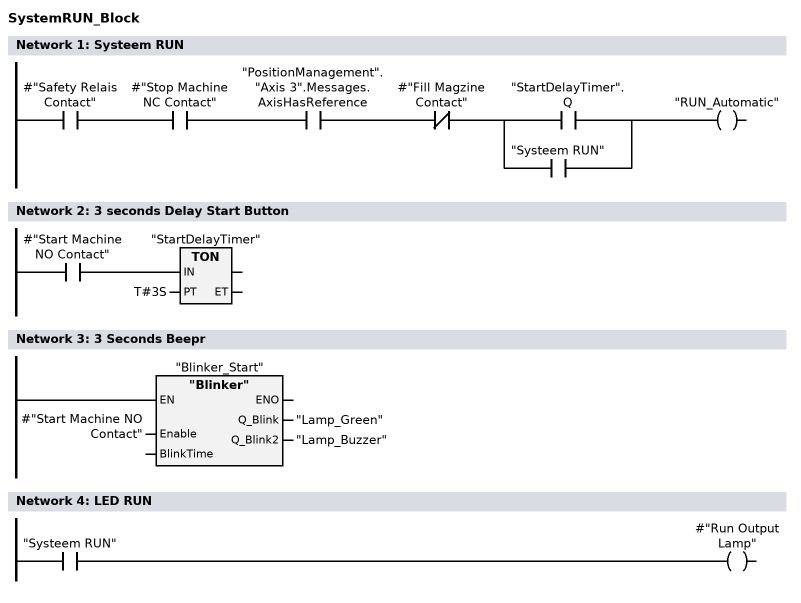
   RUNG wire#powerrail
      Contact( #"Safety Relais Contact" )
      Contact( #"Stop Machine NC Contact" )
      Contact( "PositionManagement"."Axis 3".Messages.AxisHasReference )
      I_Contact( #"Fill Magzine Contact" )
      wire#w1
      Contact( "StartDelayTimer".Q )
      wire#w2
      Coil( "RUN_Automatic" )
   END_RUNG
   RUNG wire#w1
      Contact( "Systeem RUN" )
   END_RUNG wire#w2
   // the same network as SCL:
   "RUN_Automatic" := #"Safety Relais Contact" AND #"Stop Machine NC Contact" AND "PositionManagement"."Axis 3".Messages.AxisHasReference AND NOT #"Fill Magzine Contact" AND ("StartDelayTimer".Q OR "Systeem RUN");
END_REGION

REGION Network 2: 3 seconds Delay Start Button
   "StartDelayTimer".TON(IN := #"Start Machine NO Contact", PT := T#3S);
END_REGION

REGION Network 3: 3 Seconds Beepr
   RUNG wire#powerrail
      "Blinker_Start"(Enable := #"Start Machine NO Contact", BlinkTime :=, Q_Blink => "Lamp_Green", Q_Blink2 => "Lamp_Buzzer")
   END_RUNG
   // the same network as SCL:
   "Blinker_Start"(Enable := #"Start Machine NO Contact", Q_Blink => "Lamp_Green", Q_Blink2 => "Lamp_Buzzer");   // "Blinker"
END_REGION

REGION Network 4: LED RUN
   RUNG wire#powerrail
      Contact( "Systeem RUN" )
      Coil( #"Run Output Lamp" )
   END_RUNG
   // the same network as SCL:
   #"Run Output Lamp" := "Systeem RUN";
END_REGION
END_FUNCTION

FUNCTION "SiemensEnc" : Void   // FC15, STL
TITLE = Test Siemens ENCODER
{ S7_Optimized_Access := 'FALSE' }
VERSION : 0.1
BEGIN

REGION Network 1: Presettings
         L     0;  //Delete control bits
         T     %DB1.DBD0;
         T     %DB1.DBD4;
         SET;
         S     %DB1.DBX4.0;  //Open SW gate
END_REGION

REGION Network 2: Write to the control interface
END_REGION

REGION Network 3: Read from the feedback interface
   //Read 8 bytes from the 1 Count24V
   //Configured start address of inputs
         L     "Tag_25":P;
         T     %DB1.DBD8;
         L     "Tag_26":P;
         T     %DB1.DBD12;
         R     %DB1.DBX4.0;  //Close SW gate
END_REGION
END_FUNCTION

// folder: Motion

FUNCTION_BLOCK "MC_Move"   // FB10, FBD
TITLE = MC_Move
{ S7_Optimized_Access := 'FALSE' }